HMI tags "xAO"
   "AOx_DB_M1_SP_SP" : Real = PLC AOx_DB.M1_SP.SP AT %DB203.DBD0, 1 s
   "AOx_DB_M1_SP_Signal" : Int = PLC AOx_DB.M1_SP.Signal AT %DB203.DBW6, 1 s
   "AOx_DB_M1_SP_CMD_Hand" : Bool = PLC AOx_DB.M1_SP.CMD.Hand AT %DB203.DBX8.0, 1 s
   "AOx_DB_M1_SP_CMD_Start_A" : Bool = PLC AOx_DB.M1_SP.CMD.Start_A AT %DB203.DBX8.1, 1 s
   "AOx_DB_M1_SP_CMD_Start_M" : Bool = PLC AOx_DB.M1_SP.CMD.Start_M AT %DB203.DBX8.2, 1 s
   "AOx_DB_M1_SP_SP_M" : Real = PLC AOx_DB.M1_SP.SP_M AT %DB203.DBD24, 1 s
   "AOx_DB_M1_SP_Converter_Min_In" : Real = PLC AOx_DB.M1_SP.Converter.Min_In AT %DB203.DBD46, 1 s
   "AOx_DB_M1_SP_Converter_Max_In" : Real = PLC AOx_DB.M1_SP.Converter.Max_In AT %DB203.DBD50, 1 s
   "AOx_DB_M1_SP_Converter_Min_Out" : Real = PLC AOx_DB.M1_SP.Converter.Min_Out AT %DB203.DBD54, 1 s
   "AOx_DB_M1_SP_Converter_Max_Out" : Real = PLC AOx_DB.M1_SP.Converter.Max_Out AT %DB203.DBD58, 1 s
   "AOx_DB_M2_SP_SP" : Real = PLC AOx_DB.M2_SP.SP AT %DB203.DBD98, 1 s
   "AOx_DB_M2_SP_Signal" : Int = PLC AOx_DB.M2_SP.Signal AT %DB203.DBW104, 1 s
   "AOx_DB_M2_SP_CMD_Hand" : Bool = PLC AOx_DB.M2_SP.CMD.Hand AT %DB203.DBX106.0, 1 s
   "AOx_DB_M2_SP_CMD_Start_A" : Bool = PLC AOx_DB.M2_SP.CMD.Start_A AT %DB203.DBX106.1, 1 s
   "AOx_DB_M2_SP_CMD_Start_M" : Bool = PLC AOx_DB.M2_SP.CMD.Start_M AT %DB203.DBX106.2, 1 s
   "AOx_DB_M2_SP_SP_M" : Real = PLC AOx_DB.M2_SP.SP_M AT %DB203.DBD122, 1 s
   "AOx_DB_M2_SP_Converter_Min_In" : Real = PLC AOx_DB.M2_SP.Converter.Min_In AT %DB203.DBD144, 1 s
   "AOx_DB_M2_SP_Converter_Max_In" : Real = PLC AOx_DB.M2_SP.Converter.Max_In AT %DB203.DBD148, 1 s
   "AOx_DB_M2_SP_Converter_Min_Out" : Real = PLC AOx_DB.M2_SP.Converter.Min_Out AT %DB203.DBD152, 1 s
   "AOx_DB_M2_SP_Converter_Max_Out" : Real = PLC AOx_DB.M2_SP.Converter.Max_Out AT %DB203.DBD156, 1 s
   "AOx_DB_M3_SP_SP" : Real = PLC AOx_DB.M3_SP.SP AT %DB203.DBD196, 1 s
   "AOx_DB_M3_SP_Signal" : Int = PLC AOx_DB.M3_SP.Signal AT %DB203.DBW202, 1 s
   "AOx_DB_M3_SP_CMD_Hand" : Bool = PLC AOx_DB.M3_SP.CMD.Hand AT %DB203.DBX204.0, 1 s
   "AOx_DB_M3_SP_CMD_Start_A" : Bool = PLC AOx_DB.M3_SP.CMD.Start_A AT %DB203.DBX204.1, 1 s
   "AOx_DB_M3_SP_CMD_Start_M" : Bool = PLC AOx_DB.M3_SP.CMD.Start_M AT %DB203.DBX204.2, 1 s
   "AOx_DB_M3_SP_SP_M" : Real = PLC AOx_DB.M3_SP.SP_M AT %DB203.DBD220, 1 s
   "AOx_DB_M3_SP_Converter_Min_In" : Real = PLC AOx_DB.M3_SP.Converter.Min_In AT %DB203.DBD242, 1 s
   "AOx_DB_M3_SP_Converter_Max_In" : Real = PLC AOx_DB.M3_SP.Converter.Max_In AT %DB203.DBD246, 1 s
   "AOx_DB_M3_SP_Converter_Min_Out" : Real = PLC AOx_DB.M3_SP.Converter.Min_Out AT %DB203.DBD250, 1 s
   "AOx_DB_M3_SP_Converter_Max_Out" : Real = PLC AOx_DB.M3_SP.Converter.Max_Out AT %DB203.DBD254, 1 s

HMI tags "Points"
   "Ponts_1_DB_Value" : Real = PLC Ponts_1_DB.Value AT %DB8.DBD2, 1 s
   "Ponts_1_DB_REQ" : Real = PLC Ponts_1_DB.REQ AT %DB8.DBD6, 1 s
   "Ponts_1_DB_Min" : Real = PLC Ponts_1_DB.Min AT %DB8.DBD10, 1 s
   "Ponts_1_DB_Max" : Real = PLC Ponts_1_DB.Max AT %DB8.DBD14, 1 s
   "Ponts_1_DB_SP" : Real = PLC Ponts_1_DB.SP AT %DB8.DBD18, 1 s
   "Ponts_1_DB_Now{0}" : Bool = PLC Ponts_1_DB.Now[0] AT %DB8.DBX22.0, 1 s
   "Ponts_1_DB_Now{1}" : Bool = PLC Ponts_1_DB.Now[1] AT %DB8.DBX22.1, 1 s
   "Ponts_1_DB_Now{2}" : Bool = PLC Ponts_1_DB.Now[2] AT %DB8.DBX22.2, 1 s
   "Ponts_1_DB_Now{3}" : Bool = PLC Ponts_1_DB.Now[3] AT %DB8.DBX22.3, 1 s
   "Ponts_1_DB_Now{4}" : Bool = PLC Ponts_1_DB.Now[4] AT %DB8.DBX22.4, 1 s
   "Ponts_1_DB_Now{5}" : Bool = PLC Ponts_1_DB.Now[5] AT %DB8.DBX22.5, 1 s
   "Ponts_1_DB_Now{6}" : Bool = PLC Ponts_1_DB.Now[6] AT %DB8.DBX22.6, 1 s
   "Ponts_1_DB_Now{7}" : Bool = PLC Ponts_1_DB.Now[7] AT %DB8.DBX22.7, 1 s
   "Ponts_1_DB_PLF_0_Use" : Bool = PLC Ponts_1_DB.PLF_0.Use AT %DB8.DBX24.0, 1 s
   "Ponts_1_DB_PLF_0_Low" : Real = PLC Ponts_1_DB.PLF_0.Low AT %DB8.DBD26, 1 s
   "Ponts_1_DB_PLF_0_High" : Real = PLC Ponts_1_DB.PLF_0.High AT %DB8.DBD30, 1 s
   "Ponts_1_DB_PLF_0_Point_A" : Real = PLC Ponts_1_DB.PLF_0.Point_A AT %DB8.DBD34, 1 s
   "Ponts_1_DB_PLF_0_Point_B" : Real = PLC Ponts_1_DB.PLF_0.Point_B AT %DB8.DBD38, 1 s
   "Ponts_1_DB_PLF_1_Use" : Bool = PLC Ponts_1_DB.PLF_1.Use AT %DB8.DBX44.0, 1 s
   "Ponts_1_DB_PLF_1_Low" : Real = PLC Ponts_1_DB.PLF_1.Low AT %DB8.DBD46, 1 s
   "Ponts_1_DB_PLF_1_High" : Real = PLC Ponts_1_DB.PLF_1.High AT %DB8.DBD50, 1 s
   "Ponts_1_DB_PLF_1_Point_A" : Real = PLC Ponts_1_DB.PLF_1.Point_A AT %DB8.DBD54, 1 s
   "Ponts_1_DB_PLF_1_Point_B" : Real = PLC Ponts_1_DB.PLF_1.Point_B AT %DB8.DBD58, 1 s
   "Ponts_1_DB_PLF_2_Use" : Bool = PLC Ponts_1_DB.PLF_2.Use AT %DB8.DBX64.0, 1 s
   "Ponts_1_DB_PLF_2_Low" : Real = PLC Ponts_1_DB.PLF_2.Low AT %DB8.DBD66, 1 s
   "Ponts_1_DB_PLF_2_High" : Real = PLC Ponts_1_DB.PLF_2.High AT %DB8.DBD70, 1 s
   "Ponts_1_DB_PLF_2_Point_A" : Real = PLC Ponts_1_DB.PLF_2.Point_A AT %DB8.DBD74, 1 s
   "Ponts_1_DB_PLF_2_Point_B" : Real = PLC Ponts_1_DB.PLF_2.Point_B AT %DB8.DBD78, 1 s
   "Ponts_1_DB_PLF_3_Use" : Bool = PLC Ponts_1_DB.PLF_3.Use AT %DB8.DBX84.0, 1 s
   "Ponts_1_DB_PLF_3_Low" : Real = PLC Ponts_1_DB.PLF_3.Low AT %DB8.DBD86, 1 s
   "Ponts_1_DB_PLF_3_High" : Real = PLC Ponts_1_DB.PLF_3.High AT %DB8.DBD90, 1 s
   "Ponts_1_DB_PLF_3_Point_A" : Real = PLC Ponts_1_DB.PLF_3.Point_A AT %DB8.DBD94, 1 s
   "Ponts_1_DB_PLF_3_Point_B" : Real = PLC Ponts_1_DB.PLF_3.Point_B AT %DB8.DBD98, 1 s
   "Ponts_1_DB_PLF_4_Use" : Bool = PLC Ponts_1_DB.PLF_4.Use AT %DB8.DBX104.0, 1 s
   "Ponts_1_DB_PLF_4_Low" : Real = PLC Ponts_1_DB.PLF_4.Low AT %DB8.DBD106, 1 s
   "Ponts_1_DB_PLF_4_High" : Real = PLC Ponts_1_DB.PLF_4.High AT %DB8.DBD110, 1 s
   "Ponts_1_DB_PLF_4_Point_A" : Real = PLC Ponts_1_DB.PLF_4.Point_A AT %DB8.DBD114, 1 s
   "Ponts_1_DB_PLF_4_Point_B" : Real = PLC Ponts_1_DB.PLF_4.Point_B AT %DB8.DBD118, 1 s
   "Ponts_1_DB_PLF_5_Use" : Bool = PLC Ponts_1_DB.PLF_5.Use AT %DB8.DBX124.0, 1 s
   "Ponts_1_DB_PLF_5_Low" : Real = PLC Ponts_1_DB.PLF_5.Low AT %DB8.DBD126, 1 s
   "Ponts_1_DB_PLF_5_High" : Real = PLC Ponts_1_DB.PLF_5.High AT %DB8.DBD130, 1 s
   "Ponts_1_DB_PLF_5_Point_A" : Real = PLC Ponts_1_DB.PLF_5.Point_A AT %DB8.DBD134, 1 s
   "Ponts_1_DB_PLF_5_Point_B" : Real = PLC Ponts_1_DB.PLF_5.Point_B AT %DB8.DBD138, 1 s
   "Ponts_1_DB_PLF_6_Use" : Bool = PLC Ponts_1_DB.PLF_6.Use AT %DB8.DBX144.0, 1 s
   "Ponts_1_DB_PLF_6_Low" : Real = PLC Ponts_1_DB.PLF_6.Low AT %DB8.DBD146, 1 s
   "Ponts_1_DB_PLF_6_High" : Real = PLC Ponts_1_DB.PLF_6.High AT %DB8.DBD150, 1 s
   "Ponts_1_DB_PLF_6_Point_A" : Real = PLC Ponts_1_DB.PLF_6.Point_A AT %DB8.DBD154, 1 s
   "Ponts_1_DB_PLF_6_Point_B" : Real = PLC Ponts_1_DB.PLF_6.Point_B AT %DB8.DBD158, 1 s
   "Ponts_1_DB_PLF_7_Use" : Bool = PLC Ponts_1_DB.PLF_7.Use AT %DB8.DBX164.0, 1 s
   "Ponts_1_DB_PLF_7_Low" : Real = PLC Ponts_1_DB.PLF_7.Low AT %DB8.DBD166, 1 s
   "Ponts_1_DB_PLF_7_High" : Real = PLC Ponts_1_DB.PLF_7.High AT %DB8.DBD170, 1 s
   "Ponts_1_DB_PLF_7_Point_A" : Real = PLC Ponts_1_DB.PLF_7.Point_A AT %DB8.DBD174, 1 s
   "Ponts_1_DB_PLF_7_Point_B" : Real = PLC Ponts_1_DB.PLF_7.Point_B AT %DB8.DBD178, 1 s
   "Ponts_2_DB_Value" : Real = PLC Ponts_2_DB.Value AT %DB9.DBD2, 1 s
   "Ponts_2_DB_Start" : Bool = PLC Ponts_2_DB.Start AT %DB9.DBX0.0, 1 s
   "Ponts_2_DB_REQ" : Real = PLC Ponts_2_DB.REQ AT %DB9.DBD6, 1 s
   "Ponts_2_DB_Min" : Real = PLC Ponts_2_DB.Min AT %DB9.DBD10, 1 s
   "Ponts_2_DB_Max" : Real = PLC Ponts_2_DB.Max AT %DB9.DBD14, 1 s
   "Ponts_2_DB_SP" : Real = PLC Ponts_2_DB.SP AT %DB9.DBD18, 1 s
   "Ponts_2_DB_Now{0}" : Bool = PLC Ponts_2_DB.Now[0] AT %DB9.DBX22.0, 1 s
   "Ponts_2_DB_Now{1}" : Bool = PLC Ponts_2_DB.Now[1] AT %DB9.DBX22.1, 1 s
   "Ponts_2_DB_Now{2}" : Bool = PLC Ponts_2_DB.Now[2] AT %DB9.DBX22.2, 1 s
   "Ponts_2_DB_Now{3}" : Bool = PLC Ponts_2_DB.Now[3] AT %DB9.DBX22.3, 1 s
   "Ponts_2_DB_Now{4}" : Bool = PLC Ponts_2_DB.Now[4] AT %DB9.DBX22.4, 1 s
   "Ponts_2_DB_Now{5}" : Bool = PLC Ponts_2_DB.Now[5] AT %DB9.DBX22.5, 1 s
   "Ponts_2_DB_Now{6}" : Bool = PLC Ponts_2_DB.Now[6] AT %DB9.DBX22.6, 1 s
   "Ponts_2_DB_Now{7}" : Bool = PLC Ponts_2_DB.Now[7] AT %DB9.DBX22.7, 1 s
   "Ponts_2_DB_PLF_0_Use" : Bool = PLC Ponts_2_DB.PLF_0.Use AT %DB9.DBX24.0, 1 s
   "Ponts_2_DB_PLF_0_Low" : Real = PLC Ponts_2_DB.PLF_0.Low AT %DB9.DBD26, 1 s
   "Ponts_2_DB_PLF_0_High" : Real = PLC Ponts_2_DB.PLF_0.High AT %DB9.DBD30, 1 s
   "Ponts_2_DB_PLF_0_Point_A" : Real = PLC Ponts_2_DB.PLF_0.Point_A AT %DB9.DBD34, 1 s
   "Ponts_2_DB_PLF_0_Point_B" : Real = PLC Ponts_2_DB.PLF_0.Point_B AT %DB9.DBD38, 1 s
   "Ponts_2_DB_PLF_1_Use" : Bool = PLC Ponts_2_DB.PLF_1.Use AT %DB9.DBX44.0, 1 s
   "Ponts_2_DB_PLF_1_Low" : Real = PLC Ponts_2_DB.PLF_1.Low AT %DB9.DBD46, 1 s
   "Ponts_2_DB_PLF_1_High" : Real = PLC Ponts_2_DB.PLF_1.High AT %DB9.DBD50, 1 s
   "Ponts_2_DB_PLF_1_Point_A" : Real = PLC Ponts_2_DB.PLF_1.Point_A AT %DB9.DBD54, 1 s
   "Ponts_2_DB_PLF_1_Point_B" : Real = PLC Ponts_2_DB.PLF_1.Point_B AT %DB9.DBD58, 1 s
   "Ponts_2_DB_PLF_2_Use" : Bool = PLC Ponts_2_DB.PLF_2.Use AT %DB9.DBX64.0, 1 s
   "Ponts_2_DB_PLF_2_Low" : Real = PLC Ponts_2_DB.PLF_2.Low AT %DB9.DBD66, 1 s
   "Ponts_2_DB_PLF_2_High" : Real = PLC Ponts_2_DB.PLF_2.High AT %DB9.DBD70, 1 s
   "Ponts_2_DB_PLF_2_Point_A" : Real = PLC Ponts_2_DB.PLF_2.Point_A AT %DB9.DBD74, 1 s
   "Ponts_2_DB_PLF_2_Point_B" : Real = PLC Ponts_2_DB.PLF_2.Point_B AT %DB9.DBD78, 1 s
   "Ponts_2_DB_PLF_3_Use" : Bool = PLC Ponts_2_DB.PLF_3.Use AT %DB9.DBX84.0, 1 s
   "Ponts_2_DB_PLF_3_Low" : Real = PLC Ponts_2_DB.PLF_3.Low AT %DB9.DBD86, 1 s
   "Ponts_2_DB_PLF_3_High" : Real = PLC Ponts_2_DB.PLF_3.High AT %DB9.DBD90, 1 s
   "Ponts_2_DB_PLF_3_Point_A" : Real = PLC Ponts_2_DB.PLF_3.Point_A AT %DB9.DBD94, 1 s
   "Ponts_2_DB_PLF_3_Point_B" : Real = PLC Ponts_2_DB.PLF_3.Point_B AT %DB9.DBD98, 1 s
   "Ponts_2_DB_PLF_4_Use" : Bool = PLC Ponts_2_DB.PLF_4.Use AT %DB9.DBX104.0, 1 s
   "Ponts_2_DB_PLF_4_Low" : Real = PLC Ponts_2_DB.PLF_4.Low AT %DB9.DBD106, 1 s
   "Ponts_2_DB_PLF_4_High" : Real = PLC Ponts_2_DB.PLF_4.High AT %DB9.DBD110, 1 s
   "Ponts_2_DB_PLF_4_Point_A" : Real = PLC Ponts_2_DB.PLF_4.Point_A AT %DB9.DBD114, 1 s
   "Ponts_2_DB_PLF_4_Point_B" : Real = PLC Ponts_2_DB.PLF_4.Point_B AT %DB9.DBD118, 1 s
   "Ponts_2_DB_PLF_5_Use" : Bool = PLC Ponts_2_DB.PLF_5.Use AT %DB9.DBX124.0, 1 s
   "Ponts_2_DB_PLF_5_Low" : Real = PLC Ponts_2_DB.PLF_5.Low AT %DB9.DBD126, 1 s
   "Ponts_2_DB_PLF_5_High" : Real = PLC Ponts_2_DB.PLF_5.High AT %DB9.DBD130, 1 s
   "Ponts_2_DB_PLF_5_Point_A" : Real = PLC Ponts_2_DB.PLF_5.Point_A AT %DB9.DBD134, 1 s
   "Ponts_2_DB_PLF_5_Point_B" : Real = PLC Ponts_2_DB.PLF_5.Point_B AT %DB9.DBD138, 1 s
   "Ponts_2_DB_PLF_6_Use" : Bool = PLC Ponts_2_DB.PLF_6.Use AT %DB9.DBX144.0, 1 s
   "Ponts_2_DB_PLF_6_Low" : Real = PLC Ponts_2_DB.PLF_6.Low AT %DB9.DBD146, 1 s
   "Ponts_2_DB_PLF_6_High" : Real = PLC Ponts_2_DB.PLF_6.High AT %DB9.DBD150, 1 s
   "Ponts_2_DB_PLF_6_Point_A" : Real = PLC Ponts_2_DB.PLF_6.Point_A AT %DB9.DBD154, 1 s
   "Ponts_2_DB_PLF_6_Point_B" : Real = PLC Ponts_2_DB.PLF_6.Point_B AT %DB9.DBD158, 1 s
   "Ponts_2_DB_PLF_7_Use" : Bool = PLC Ponts_2_DB.PLF_7.Use AT %DB9.DBX164.0, 1 s
   "Ponts_2_DB_PLF_7_Low" : Real = PLC Ponts_2_DB.PLF_7.Low AT %DB9.DBD166, 1 s
   "Ponts_2_DB_PLF_7_High" : Real = PLC Ponts_2_DB.PLF_7.High AT %DB9.DBD170, 1 s
   "Ponts_2_DB_PLF_7_Point_A" : Real = PLC Ponts_2_DB.PLF_7.Point_A AT %DB9.DBD174, 1 s
   "Ponts_2_DB_PLF_7_Point_B" : Real = PLC Ponts_2_DB.PLF_7.Point_B AT %DB9.DBD178, 1 s

HMI tags "Mass"
   "Statistics_DB_Summ_1" : Real = PLC Statistics_DB.Summ_1 AT %DB4.DBD48, 1 s
   "Statistics_DB_Summ_2" : Real = PLC Statistics_DB.Summ_2 AT %DB4.DBD52, 1 s
   "Statistics_DB_All_1" : Real = PLC Statistics_DB.All_1 AT %DB4.DBD56, 1 s
   "Statistics_DB_All_2" : Real = PLC Statistics_DB.All_2 AT %DB4.DBD60, 1 s
   "Statistics_DB_Last_Month_1" : Real = PLC Statistics_DB.Last_Month_1 AT %DB4.DBD572, 1 s
   "Statistics_DB_Last_Month_2" : Real = PLC Statistics_DB.Last_Month_2 AT %DB4.DBD576, 1 s
   "Statistics_DB_Month_1{1}" : Real = PLC Statistics_DB.Month_1[1] AT %DB4.DBD76, 1 s
   "Statistics_DB_Month_1{2}" : Real = PLC Statistics_DB.Month_1[2] AT %DB4.DBD80, 1 s
   "Statistics_DB_Month_1{3}" : Real = PLC Statistics_DB.Month_1[3] AT %DB4.DBD84, 1 s
   "Statistics_DB_Month_1{4}" : Real = PLC Statistics_DB.Month_1[4] AT %DB4.DBD88, 1 s
   "Statistics_DB_Month_1{5}" : Real = PLC Statistics_DB.Month_1[5] AT %DB4.DBD92, 1 s
   "Statistics_DB_Month_1{6}" : Real = PLC Statistics_DB.Month_1[6] AT %DB4.DBD96, 1 s
   "Statistics_DB_Month_1{7}" : Real = PLC Statistics_DB.Month_1[7] AT %DB4.DBD100, 1 s
   "Statistics_DB_Month_1{8}" : Real = PLC Statistics_DB.Month_1[8] AT %DB4.DBD104, 1 s
   "Statistics_DB_Month_1{9}" : Real = PLC Statistics_DB.Month_1[9] AT %DB4.DBD108, 1 s
   "Statistics_DB_Month_1{10}" : Real = PLC Statistics_DB.Month_1[10] AT %DB4.DBD112, 1 s
   "Statistics_DB_Month_1{11}" : Real = PLC Statistics_DB.Month_1[11] AT %DB4.DBD116, 1 s
   "Statistics_DB_Month_1{12}" : Real = PLC Statistics_DB.Month_1[12] AT %DB4.DBD120, 1 s
   "Statistics_DB_Month_1{13}" : Real = PLC Statistics_DB.Month_1[13] AT %DB4.DBD124, 1 s
   "Statistics_DB_Month_1{14}" : Real = PLC Statistics_DB.Month_1[14] AT %DB4.DBD128, 1 s
   "Statistics_DB_Month_1{15}" : Real = PLC Statistics_DB.Month_1[15] AT %DB4.DBD132, 1 s
   "Statistics_DB_Month_1{16}" : Real = PLC Statistics_DB.Month_1[16] AT %DB4.DBD136, 1 s
   "Statistics_DB_Month_1{17}" : Real = PLC Statistics_DB.Month_1[17] AT %DB4.DBD140, 1 s
   "Statistics_DB_Month_1{18}" : Real = PLC Statistics_DB.Month_1[18] AT %DB4.DBD144, 1 s
   "Statistics_DB_Month_1{19}" : Real = PLC Statistics_DB.Month_1[19] AT %DB4.DBD148, 1 s
   "Statistics_DB_Month_1{20}" : Real = PLC Statistics_DB.Month_1[20] AT %DB4.DBD152, 1 s
   "Statistics_DB_Month_1{21}" : Real = PLC Statistics_DB.Month_1[21] AT %DB4.DBD156, 1 s
   "Statistics_DB_Month_1{22}" : Real = PLC Statistics_DB.Month_1[22] AT %DB4.DBD160, 1 s
   "Statistics_DB_Month_1{23}" : Real = PLC Statistics_DB.Month_1[23] AT %DB4.DBD164, 1 s
   "Statistics_DB_Month_1{24}" : Real = PLC Statistics_DB.Month_1[24] AT %DB4.DBD168, 1 s
   "Statistics_DB_Month_1{25}" : Real = PLC Statistics_DB.Month_1[25] AT %DB4.DBD172, 1 s
   "Statistics_DB_Month_1{26}" : Real = PLC Statistics_DB.Month_1[26] AT %DB4.DBD176, 1 s
   "Statistics_DB_Month_1{27}" : Real = PLC Statistics_DB.Month_1[27] AT %DB4.DBD180, 1 s
   "Statistics_DB_Month_1{28}" : Real = PLC Statistics_DB.Month_1[28] AT %DB4.DBD184, 1 s
   "Statistics_DB_Month_1{29}" : Real = PLC Statistics_DB.Month_1[29] AT %DB4.DBD188, 1 s
   "Statistics_DB_Month_1{30}" : Real = PLC Statistics_DB.Month_1[30] AT %DB4.DBD192, 1 s
   "Statistics_DB_Month_1{31}" : Real = PLC Statistics_DB.Month_1[31] AT %DB4.DBD196, 1 s
   "Statistics_DB_Month_2{1}" : Real = PLC Statistics_DB.Month_2[1] AT %DB4.DBD200, 1 s
   "Statistics_DB_Month_2{2}" : Real = PLC Statistics_DB.Month_2[2] AT %DB4.DBD204, 1 s
   "Statistics_DB_Month_2{3}" : Real = PLC Statistics_DB.Month_2[3] AT %DB4.DBD208, 1 s
   "Statistics_DB_Month_2{4}" : Real = PLC Statistics_DB.Month_2[4] AT %DB4.DBD212, 1 s
   "Statistics_DB_Month_2{5}" : Real = PLC Statistics_DB.Month_2[5] AT %DB4.DBD216, 1 s
   "Statistics_DB_Month_2{6}" : Real = PLC Statistics_DB.Month_2[6] AT %DB4.DBD220, 1 s
   "Statistics_DB_Month_2{7}" : Real = PLC Statistics_DB.Month_2[7] AT %DB4.DBD224, 1 s
   "Statistics_DB_Month_2{8}" : Real = PLC Statistics_DB.Month_2[8] AT %DB4.DBD228, 1 s
   "Statistics_DB_Month_2{9}" : Real = PLC Statistics_DB.Month_2[9] AT %DB4.DBD232, 1 s
   "Statistics_DB_Month_2{10}" : Real = PLC Statistics_DB.Month_2[10] AT %DB4.DBD236, 1 s
   "Statistics_DB_Month_2{11}" : Real = PLC Statistics_DB.Month_2[11] AT %DB4.DBD240, 1 s
   "Statistics_DB_Month_2{12}" : Real = PLC Statistics_DB.Month_2[12] AT %DB4.DBD244, 1 s
   "Statistics_DB_Month_2{13}" : Real = PLC Statistics_DB.Month_2[13] AT %DB4.DBD248, 1 s
   "Statistics_DB_Month_2{14}" : Real = PLC Statistics_DB.Month_2[14] AT %DB4.DBD252, 1 s
   "Statistics_DB_Month_2{15}" : Real = PLC Statistics_DB.Month_2[15] AT %DB4.DBD256, 1 s
   "Statistics_DB_Month_2{16}" : Real = PLC Statistics_DB.Month_2[16] AT %DB4.DBD260, 1 s
   "Statistics_DB_Month_2{17}" : Real = PLC Statistics_DB.Month_2[17] AT %DB4.DBD264, 1 s
   "Statistics_DB_Month_2{18}" : Real = PLC Statistics_DB.Month_2[18] AT %DB4.DBD268, 1 s
   "Statistics_DB_Month_2{19}" : Real = PLC Statistics_DB.Month_2[19] AT %DB4.DBD272, 1 s
   "Statistics_DB_Month_2{20}" : Real = PLC Statistics_DB.Month_2[20] AT %DB4.DBD276, 1 s
   "Statistics_DB_Month_2{21}" : Real = PLC Statistics_DB.Month_2[21] AT %DB4.DBD280, 1 s
   "Statistics_DB_Month_2{22}" : Real = PLC Statistics_DB.Month_2[22] AT %DB4.DBD284, 1 s
   "Statistics_DB_Month_2{23}" : Real = PLC Statistics_DB.Month_2[23] AT %DB4.DBD288, 1 s
   "Statistics_DB_Month_2{24}" : Real = PLC Statistics_DB.Month_2[24] AT %DB4.DBD292, 1 s
   "Statistics_DB_Month_2{25}" : Real = PLC Statistics_DB.Month_2[25] AT %DB4.DBD296, 1 s
   "Statistics_DB_Month_2{26}" : Real = PLC Statistics_DB.Month_2[26] AT %DB4.DBD300, 1 s
   "Statistics_DB_Month_2{27}" : Real = PLC Statistics_DB.Month_2[27] AT %DB4.DBD304, 1 s
   "Statistics_DB_Month_2{28}" : Real = PLC Statistics_DB.Month_2[28] AT %DB4.DBD308, 1 s
   "Statistics_DB_Month_2{29}" : Real = PLC Statistics_DB.Month_2[29] AT %DB4.DBD312, 1 s
   "Statistics_DB_Month_2{30}" : Real = PLC Statistics_DB.Month_2[30] AT %DB4.DBD316, 1 s
   "Statistics_DB_Month_2{31}" : Real = PLC Statistics_DB.Month_2[31] AT %DB4.DBD320, 1 s
   "Statistics_DB_Last_M_1{1}" : Real = PLC Statistics_DB.Last_M_1[1] AT %DB4.DBD324, 1 s
   "Statistics_DB_Last_M_1{2}" : Real = PLC Statistics_DB.Last_M_1[2] AT %DB4.DBD328, 1 s
   "Statistics_DB_Last_M_1{3}" : Real = PLC Statistics_DB.Last_M_1[3] AT %DB4.DBD332, 1 s
   "Statistics_DB_Last_M_1{4}" : Real = PLC Statistics_DB.Last_M_1[4] AT %DB4.DBD336, 1 s
   "Statistics_DB_Last_M_1{5}" : Real = PLC Statistics_DB.Last_M_1[5] AT %DB4.DBD340, 1 s
   "Statistics_DB_Last_M_1{6}" : Real = PLC Statistics_DB.Last_M_1[6] AT %DB4.DBD344, 1 s
   "Statistics_DB_Last_M_1{7}" : Real = PLC Statistics_DB.Last_M_1[7] AT %DB4.DBD348, 1 s
   "Statistics_DB_Last_M_1{8}" : Real = PLC Statistics_DB.Last_M_1[8] AT %DB4.DBD352, 1 s
   "Statistics_DB_Last_M_1{9}" : Real = PLC Statistics_DB.Last_M_1[9] AT %DB4.DBD356, 1 s
   "Statistics_DB_Last_M_1{10}" : Real = PLC Statistics_DB.Last_M_1[10] AT %DB4.DBD360, 1 s
   "Statistics_DB_Last_M_1{11}" : Real = PLC Statistics_DB.Last_M_1[11] AT %DB4.DBD364, 1 s
   "Statistics_DB_Last_M_1{12}" : Real = PLC Statistics_DB.Last_M_1[12] AT %DB4.DBD368, 1 s
   "Statistics_DB_Last_M_1{13}" : Real = PLC Statistics_DB.Last_M_1[13] AT %DB4.DBD372, 1 s
   "Statistics_DB_Last_M_1{14}" : Real = PLC Statistics_DB.Last_M_1[14] AT %DB4.DBD376, 1 s
   "Statistics_DB_Last_M_1{15}" : Real = PLC Statistics_DB.Last_M_1[15] AT %DB4.DBD380, 1 s
   "Statistics_DB_Last_M_1{16}" : Real = PLC Statistics_DB.Last_M_1[16] AT %DB4.DBD384, 1 s
   "Statistics_DB_Last_M_1{17}" : Real = PLC Statistics_DB.Last_M_1[17] AT %DB4.DBD388, 1 s
   "Statistics_DB_Last_M_1{18}" : Real = PLC Statistics_DB.Last_M_1[18] AT %DB4.DBD392, 1 s
   "Statistics_DB_Last_M_1{19}" : Real = PLC Statistics_DB.Last_M_1[19] AT %DB4.DBD396, 1 s
   "Statistics_DB_Last_M_1{20}" : Real = PLC Statistics_DB.Last_M_1[20] AT %DB4.DBD400, 1 s
   "Statistics_DB_Last_M_1{21}" : Real = PLC Statistics_DB.Last_M_1[21] AT %DB4.DBD404, 1 s
   "Statistics_DB_Last_M_1{22}" : Real = PLC Statistics_DB.Last_M_1[22] AT %DB4.DBD408, 1 s
   "Statistics_DB_Last_M_1{23}" : Real = PLC Statistics_DB.Last_M_1[23] AT %DB4.DBD412, 1 s
   "Statistics_DB_Last_M_1{24}" : Real = PLC Statistics_DB.Last_M_1[24] AT %DB4.DBD416, 1 s
   "Statistics_DB_Last_M_1{25}" : Real = PLC Statistics_DB.Last_M_1[25] AT %DB4.DBD420, 1 s
   "Statistics_DB_Last_M_1{26}" : Real = PLC Statistics_DB.Last_M_1[26] AT %DB4.DBD424, 1 s
   "Statistics_DB_Last_M_1{27}" : Real = PLC Statistics_DB.Last_M_1[27] AT %DB4.DBD428, 1 s
   "Statistics_DB_Last_M_1{28}" : Real = PLC Statistics_DB.Last_M_1[28] AT %DB4.DBD432, 1 s
   "Statistics_DB_Last_M_1{29}" : Real = PLC Statistics_DB.Last_M_1[29] AT %DB4.DBD436, 1 s
   "Statistics_DB_Last_M_1{30}" : Real = PLC Statistics_DB.Last_M_1[30] AT %DB4.DBD440, 1 s
   "Statistics_DB_Last_M_1{31}" : Real = PLC Statistics_DB.Last_M_1[31] AT %DB4.DBD444, 1 s
   "Statistics_DB_Last_M_2{1}" : Real = PLC Statistics_DB.Last_M_2[1] AT %DB4.DBD448, 1 s
   "Statistics_DB_Last_M_2{2}" : Real = PLC Statistics_DB.Last_M_2[2] AT %DB4.DBD452, 1 s
   "Statistics_DB_Last_M_2{3}" : Real = PLC Statistics_DB.Last_M_2[3] AT %DB4.DBD456, 1 s
   "Statistics_DB_Last_M_2{4}" : Real = PLC Statistics_DB.Last_M_2[4] AT %DB4.DBD460, 1 s
   "Statistics_DB_Last_M_2{5}" : Real = PLC Statistics_DB.Last_M_2[5] AT %DB4.DBD464, 1 s
   "Statistics_DB_Last_M_2{6}" : Real = PLC Statistics_DB.Last_M_2[6] AT %DB4.DBD468, 1 s
   "Statistics_DB_Last_M_2{7}" : Real = PLC Statistics_DB.Last_M_2[7] AT %DB4.DBD472, 1 s
   "Statistics_DB_Last_M_2{8}" : Real = PLC Statistics_DB.Last_M_2[8] AT %DB4.DBD476, 1 s
   "Statistics_DB_Last_M_2{9}" : Real = PLC Statistics_DB.Last_M_2[9] AT %DB4.DBD480, 1 s
   "Statistics_DB_Last_M_2{10}" : Real = PLC Statistics_DB.Last_M_2[10] AT %DB4.DBD484, 1 s
   "Statistics_DB_Last_M_2{11}" : Real = PLC Statistics_DB.Last_M_2[11] AT %DB4.DBD488, 1 s
   "Statistics_DB_Last_M_2{12}" : Real = PLC Statistics_DB.Last_M_2[12] AT %DB4.DBD492, 1 s
   "Statistics_DB_Last_M_2{13}" : Real = PLC Statistics_DB.Last_M_2[13] AT %DB4.DBD496, 1 s
   "Statistics_DB_Last_M_2{14}" : Real = PLC Statistics_DB.Last_M_2[14] AT %DB4.DBD500, 1 s
   "Statistics_DB_Last_M_2{15}" : Real = PLC Statistics_DB.Last_M_2[15] AT %DB4.DBD504, 1 s
   "Statistics_DB_Last_M_2{16}" : Real = PLC Statistics_DB.Last_M_2[16] AT %DB4.DBD508, 1 s
   "Statistics_DB_Last_M_2{17}" : Real = PLC Statistics_DB.Last_M_2[17] AT %DB4.DBD512, 1 s
   "Statistics_DB_Last_M_2{18}" : Real = PLC Statistics_DB.Last_M_2[18] AT %DB4.DBD516, 1 s
   "Statistics_DB_Last_M_2{19}" : Real = PLC Statistics_DB.Last_M_2[19] AT %DB4.DBD520, 1 s
   "Statistics_DB_Last_M_2{20}" : Real = PLC Statistics_DB.Last_M_2[20] AT %DB4.DBD524, 1 s
   "Statistics_DB_Last_M_2{21}" : Real = PLC Statistics_DB.Last_M_2[21] AT %DB4.DBD528, 1 s
   "Statistics_DB_Last_M_2{22}" : Real = PLC Statistics_DB.Last_M_2[22] AT %DB4.DBD532, 1 s
   "Statistics_DB_Last_M_2{23}" : Real = PLC Statistics_DB.Last_M_2[23] AT %DB4.DBD536, 1 s
   "Statistics_DB_Last_M_2{24}" : Real = PLC Statistics_DB.Last_M_2[24] AT %DB4.DBD540, 1 s
   "Statistics_DB_Last_M_2{25}" : Real = PLC Statistics_DB.Last_M_2[25] AT %DB4.DBD544, 1 s
   "Statistics_DB_Last_M_2{26}" : Real = PLC Statistics_DB.Last_M_2[26] AT %DB4.DBD548, 1 s
   "Statistics_DB_Last_M_2{27}" : Real = PLC Statistics_DB.Last_M_2[27] AT %DB4.DBD552, 1 s
   "Statistics_DB_Last_M_2{28}" : Real = PLC Statistics_DB.Last_M_2[28] AT %DB4.DBD556, 1 s
   "Statistics_DB_Last_M_2{29}" : Real = PLC Statistics_DB.Last_M_2[29] AT %DB4.DBD560, 1 s
   "Statistics_DB_Last_M_2{30}" : Real = PLC Statistics_DB.Last_M_2[30] AT %DB4.DBD564, 1 s
   "Statistics_DB_Last_M_2{31}" : Real = PLC Statistics_DB.Last_M_2[31] AT %DB4.DBD568, 1 s

HMI tags "PID"
   "PID_M1_SP" : Real = PLC PID_M1.SP AT %DB5.DBD2, 1 s
   "PID_M1_Value" : Real = PLC PID_M1.Value AT %DB5.DBD6, 1 s
   "PID_M1_Hand" : Bool = PLC PID_M1.Hand AT %DB5.DBX14.0, 1 s
   "PID_M1_Reset" : Bool = PLC PID_M1.Reset AT %DB5.DBX14.2, 1 s
   "PID_M1_Invert" : Bool = PLC PID_M1.Invert AT %DB5.DBX14.4, 1 s
   "PID_M1_HandValue" : Real = PLC PID_M1.HandValue AT %DB5.DBD24, 1 s
   "PID_M1_SP_P" : Real = PLC PID_M1.SP_P AT %DB5.DBD28, 1 s
   "PID_M1_SP_Ti" : Real = PLC PID_M1.SP_Ti AT %DB5.DBD32, 1 s
   "PID_M1_SP_Td" : Real = PLC PID_M1.SP_Td AT %DB5.DBD36, 1 s
   "PID_M1_SP_Cycle" : Real = PLC PID_M1.SP_Cycle AT %DB5.DBD40, 1 s
   "PID_M1_Max_SP" : Real = PLC PID_M1.Max_SP AT %DB5.DBD48, 1 s
   "PID_M1_Min_SP" : Real = PLC PID_M1.Min_SP AT %DB5.DBD52, 1 s
   "PID_M1_Max_in" : Real = PLC PID_M1.Max_in AT %DB5.DBD56, 1 s
   "PID_M1_Min_in" : Real = PLC PID_M1.Min_in AT %DB5.DBD60, 1 s
   "PID_M1_Max_out" : Real = PLC PID_M1.Max_out AT %DB5.DBD64, 1 s
   "PID_M1_Min_out" : Real = PLC PID_M1.Min_out AT %DB5.DBD68, 1 s
   "PID_M1_DeadBand" : Real = PLC PID_M1.DeadBand AT %DB5.DBD78, 1 s
   "PID_M1_Converter_Min_In" : Real = PLC PID_M1.Converter.Min_In AT %DB5.DBD92, 1 s
   "PID_M1_Converter_Max_In" : Real = PLC PID_M1.Converter.Max_In AT %DB5.DBD96, 1 s
   "PID_M1_Converter_Min_Out" : Real = PLC PID_M1.Converter.Min_Out AT %DB5.DBD100, 1 s
   "PID_M1_Converter_Max_Out" : Real = PLC PID_M1.Converter.Max_Out AT %DB5.DBD104, 1 s
   "PID_M2_SP" : Real = PLC PID_M2.SP AT %DB6.DBD2, 1 s
   "PID_M2_Value" : Real = PLC PID_M2.Value AT %DB6.DBD6, 1 s
   "PID_M2_Hand" : Bool = PLC PID_M2.Hand AT %DB6.DBX14.0, 1 s
   "PID_M2_Reset" : Bool = PLC PID_M2.Reset AT %DB6.DBX14.2, 1 s
   "PID_M2_Invert" : Bool = PLC PID_M2.Invert AT %DB6.DBX14.4, 1 s
   "PID_M2_HandValue" : Real = PLC PID_M2.HandValue AT %DB6.DBD24, 1 s
   "PID_M2_SP_P" : Real = PLC PID_M2.SP_P AT %DB6.DBD28, 1 s
   "PID_M2_SP_Ti" : Real = PLC PID_M2.SP_Ti AT %DB6.DBD32, 1 s
   "PID_M2_SP_Td" : Real = PLC PID_M2.SP_Td AT %DB6.DBD36, 1 s
   "PID_M2_SP_Cycle" : Real = PLC PID_M2.SP_Cycle AT %DB6.DBD40, 1 s
   "PID_M2_Max_SP" : Real = PLC PID_M2.Max_SP AT %DB6.DBD48, 1 s
   "PID_M2_Min_SP" : Real = PLC PID_M2.Min_SP AT %DB6.DBD52, 1 s
   "PID_M2_Max_in" : Real = PLC PID_M2.Max_in AT %DB6.DBD56, 1 s
   "PID_M2_Min_in" : Real = PLC PID_M2.Min_in AT %DB6.DBD60, 1 s
   "PID_M2_Max_out" : Real = PLC PID_M2.Max_out AT %DB6.DBD64, 1 s
   "PID_M2_Min_out" : Real = PLC PID_M2.Min_out AT %DB6.DBD68, 1 s
   "PID_M2_Converter_Min_In" : Real = PLC PID_M2.Converter.Min_In AT %DB6.DBD92, 1 s
   "PID_M2_Converter_Max_In" : Real = PLC PID_M2.Converter.Max_In AT %DB6.DBD96, 1 s
   "PID_M2_Converter_Min_Out" : Real = PLC PID_M2.Converter.Min_Out AT %DB6.DBD100, 1 s
   "PID_M2_Converter_Max_Out" : Real = PLC PID_M2.Converter.Max_Out AT %DB6.DBD104, 1 s
   "PID_M2_DeadBand" : Real = PLC PID_M2.DeadBand AT %DB6.DBD78, 1 s

discrete alarms
   11: 'Расходомер 1 - Обрыв датчика', class Errors, trigger "AIx_DB_Flow_1_Alarm" bit 0
   12: 'Расходомер 1 - Короткое замыкание', class Errors, trigger "AIx_DB_Flow_1_Alarm" bit 1
   13: 'Расходомер 1 - Аварийно высокий поток', class Errors, trigger "AIx_DB_Flow_1_Alarm" bit 2
   14: 'Расходомер 1 - Высокий поток', class Errors, trigger "AIx_DB_Flow_1_Alarm" bit 3
   15: 'Расходомер 1 - Низкий поток', class Errors, trigger "AIx_DB_Flow_1_Alarm" bit 4
   16: 'Расходомер 1 - Аварийно низкий поток', class Errors, trigger "AIx_DB_Flow_1_Alarm" bit 5
   17: 'Дозатор 1 - Выбило защитный автомат', class Errors, trigger "Motors_DB_M1_Alarm" bit 0
   18: 'Дозатор 1 - Ошибка при запуске', class Errors, trigger "Motors_DB_M1_Alarm" bit 1
   19: 'Дозатор 1 - Ошибка при останове', class Errors, trigger "Motors_DB_M1_Alarm" bit 2
   20: 'Дозатор 1 - Сработало реле безопасности', class Errors, trigger "Motors_DB_M1_Alarm" bit 3
   21: 'Дозатор 1 - Общая блокировка', class Errors, trigger "Motors_DB_M1_Alarm" bit 4
   22: 'Дозатор 1 - Перегрев двигателя', class Errors, trigger "Motors_DB_M1_Alarm" bit 5
   23: 'Дозатор 2 - Выбило защитный автомат', class Errors, trigger "Motors_DB_M2_Alarm" bit 0
   24: 'Дозатор 2 - Ошибка при запуске', class Errors, trigger "Motors_DB_M2_Alarm" bit 1
   25: 'Дозатор 2 - Ошибка при останове', class Errors, trigger "Motors_DB_M2_Alarm" bit 2
   26: 'Дозатор 2 - Сработало реле безопасности', class Errors, trigger "Motors_DB_M2_Alarm" bit 3
   27: 'Дозатор 2 - Общая блокировка', class Errors, trigger "Motors_DB_M2_Alarm" bit 4
   28: 'Дозатор 2 - Перегрев двигателя', class Errors, trigger "Motors_DB_M2_Alarm" bit 5
   29: 'Дозатор 3 - Выбило защитный автомат', class Errors, trigger "Motors_DB_M3_Alarm" bit 0
   30: 'Дозатор 3 - Ошибка при запуске', class Errors, trigger "Motors_DB_M3_Alarm" bit 1
   31: 'Дозатор 3 - Ошибка при останове', class Errors, trigger "Motors_DB_M3_Alarm" bit 2
   32: 'Дозатор 3 - Сработало реле безопасности', class Errors, trigger "Motors_DB_M3_Alarm" bit 3
   33: 'Дозатор 3 - Общая блокировка', class Errors, trigger "Motors_DB_M3_Alarm" bit 4
   34: 'Дозатор 3 - Перегрев двигателя', class Errors, trigger "Motors_DB_M3_Alarm" bit 5
   53: 'Расходомер 2 - Обрыв датчика', class Errors, trigger "AIx_DB_Flow_2_Alarm" bit 0
   54: 'Расходомер 2 - Короткое замыкание', class Errors, trigger "AIx_DB_Flow_2_Alarm" bit 1
   55: 'Расходомер 2 - Аварийно высокий поток', class Errors, trigger "AIx_DB_Flow_2_Alarm" bit 2
   56: 'Расходомер 2 - Высокий поток', class Errors, trigger "AIx_DB_Flow_2_Alarm" bit 3
   57: 'Расходомер 2 - Низкий поток', class Errors, trigger "AIx_DB_Flow_2_Alarm" bit 4
   58: 'Расходомер 2 - Аварийно низкий поток', class Errors, trigger "AIx_DB_Flow_2_Alarm" bit 5
   35: 'Мутность 1 - Обрыв датчика', class Errors, trigger "AIx_DB_Trans_1_Alarm" bit 0
   36: 'Мутность 1 - Короткое замыкание', class Errors, trigger "AIx_DB_Trans_1_Alarm" bit 1
   37: 'Мутность 1 - Аварийно высокий порог', class Errors, trigger "AIx_DB_Trans_1_Alarm" bit 2
   38: 'Мутность 1 - Высокий порог', class Errors, trigger "AIx_DB_Trans_1_Alarm" bit 3
   39: 'Мутность 1 - Низкий порог', class Errors, trigger "AIx_DB_Trans_1_Alarm" bit 4
   40: 'Мутность 1 - Аварийно низкий порог', class Errors, trigger "AIx_DB_Trans_1_Alarm" bit 5
   59: 'Мутность 2 - Обрыв датчика', class Errors, trigger "AIx_DB_Trans_2_Alarm" bit 0
   60: 'Мутность 2 - Короткое замыкание', class Errors, trigger "AIx_DB_Trans_2_Alarm" bit 1
   61: 'Мутность 2 - Аварийно высокий порог', class Errors, trigger "AIx_DB_Trans_2_Alarm" bit 2
   62: 'Мутность 2 - Высокий порог', class Errors, trigger "AIx_DB_Trans_2_Alarm" bit 3
   63: 'Мутность 2 - Низкий порог', class Errors, trigger "AIx_DB_Trans_2_Alarm" bit 4
   64: 'Мутность 2 - Аварийно низкий порог', class Errors, trigger "AIx_DB_Trans_2_Alarm" bit 5

text list "Hand": 0 'Авто'; 1 'Ручной'

text list "настройки": 0 'Настройки >>'; 1 'Настройки <<'

graphic list "Motor": 0 'm_off_1'; 1 'm_on_1'; 2..8 'm_wait_1'; 9..1000 'm_alarm_1'

graphic list "Pump": 0 'p_off1'; 1 'p_on1'; 2..8 'p_wait1'; 9..1000 'p_alarm1'

graphic list "Valve": 0 'v_off'; 1 'v_on'; 2..8 'v_wait'; 9..1000 'v_alarm'

graphic list "L_1": 0 'L_1_off'; 1 'L_1_on'; 2..8 'L_1_wait'; 9..1000 'L_1_alarm'

graphic list "L_2": 0 'L_2_off'; 1 'L_2_on'; 2..8 'L_2_wait'; 9..1000 'L_2_alarm'

graphic list "Led": 0 'no_alarm_led'; 1 'alarm_led'

graphic list "Alarm": 0 'no_alarm_1'; 1 'alarm'

graphic list "ON_OFF": 0 'off_toggle'; 1 'on_toggle'

graphic list "ok": 0 'check_box_off'; 1 'check_box_on'

graphic list "Status": 0 'sys_x'; 1 'sys_check-mark'; 2 'z2use'; 3..99 'alarm_on'

graphic list "Vibro": 0 'b_1'; 1 'b_4'; 2..4 'b_2'; 5..1000 'b_3'

graphic list "on_off_1": 0 'check_box_off'; 1 'check_box_on'